(* Logix 5000 project; controller MV vendor 1 type 14 code 217 rev 31.11; software revision 31.00; part 47 of 53 *)
(* tags used below, declared in another part *)
   CWD : CHECKWORD_FLAGS;
   Delphi_Does_Eng_Func : BOOL;
   MV_MV10_CV1 : PlantItem;   // MV10_CV1
   MV_MV11_CV1 : PlantItem;   // MV11_CV1
   MV_MV12_CV1 : PlantItem;   // MV12_CV1
   MV_MV13_CV1 : PlantItem;   // MV13_CV1
   MV_MV14_CV1 : PlantItem;   // MV14_CV1
   MV_MV15_CV1 : PlantItem;   // MV15_CV1
   MV_MV16_CV1 : PlantItem;   // MV16_CV1
   MV_MV17_CV1 : PlantItem;   // MV17_CV1
   MV_MV18_CV1 : PlantItem;   // MV18_CV1
   MV_MV19_CV1 : PlantItem;   // MV19_CV1
   MV_MV1_CV1 : PlantItem;   // MV1_CV1
   MV_MV2_CV1 : PlantItem;   // MV2_CV1
   MV_MV30_CV1 : PlantItem;   // MV30_CV1
   MV_MV31_CV1 : PlantItem;   // MV31_CV1
   MV_MV32_CV1 : PlantItem;   // MV32_CV1
   MV_MV33_CV1 : PlantItem;   // MV33_CV1
   MV_MV34_CV1 : PlantItem;   // MV34_CV1
   MV_MV3_CV1 : PlantItem;   // MV3_CV1
   MV_MV4_CV1 : PlantItem;   // MV4_CV1
   MV_MV5_CV1 : PlantItem;   // MV5_CV1
   MV_MV6_CV1 : PlantItem;   // MV6_CV1
   MV_MV7_CV1 : PlantItem;   // MV7_CV1
   MV_MV8_CV1 : PlantItem;   // MV8_CV1
   MV_MV9_CV1 : PlantItem;   // MV9_CV1
   MV_N255 : DINT[255];   // Old Format Checkwords To Keep Delphi Indicating Status Correctly.
(* MV_Common, continued *)

ROUTINE MV_Old_Checkword_Relaying   (* ladder *)
// Relay New Item Format To Old CW To Keep Delphi Happy Until Full Changeover.
   0: [XIC(Delphi_Does_Eng_Func) [[XIC(MV_N255[0].8) [OTL(MV_MV1_CV1.CW.[CWD.MANUAL]) ,XIC(MV_N255[0].9) OTL(MV_MV1_CV1.CW.[CWD.MANDRV]) ,XIO(MV_N255[0].9) OTU(MV_MV1_CV1.CW.[CWD.MANDRV]) ] ,XIO(MV_N255[0].8) [OTU(MV_MV1_CV1.CW.[CWD.MANUAL]) ,[XIC(MV_MV1_CV1.CW.[CWD.OUTPUT]) OTL(MV_N255[0].9) ,XIO(MV_MV1_CV1.CW.[CWD.OUTPUT]) OTU(MV_N255[0].9) ] ] ] ,[XIC(MV_N255[0].13) OTL(MV_MV1_CV1.CW.[CWD.CHECKOFF]) ,XIO(MV_N255[0].13) OTU(MV_MV1_CV1.CW.[CWD.CHECKOFF]) ] ] ,XIO(Delphi_Does_Eng_Func) [[XIC(MV_MV1_CV1.CW.[CWD.MANUAL]) OTL(MV_N255[0].8) ,XIO(MV_MV1_CV1.CW.[CWD.MANUAL]) OTU(MV_N255[0].8) ] ,[XIC(MV_MV1_CV1.CW.[CWD.CHECKOFF]) OTL(MV_N255[0].13) ,XIO(MV_MV1_CV1.CW.[CWD.CHECKOFF]) OTU(MV_N255[0].13) ] ,[XIC(MV_MV1_CV1.CW.[CWD.OUTPUT]) OTL(MV_N255[0].9) ,XIO(MV_MV1_CV1.CW.[CWD.OUTPUT]) OTU(MV_N255[0].9) ] ] ,XIC(MV_MV1_CV1.CW.[CWD.OUTPUT]) OTE(MV_N255[0].10) ,XIO(MV_MV1_CV1.CW.[CWD.OUTPUT]) OTE(MV_N255[0].11) ,XIC(MV_MV1_CV1.CW.[CWD.FAULT]) OTE(MV_N255[0].15) ];
   1: [XIC(Delphi_Does_Eng_Func) [[XIC(MV_N255[1].8) [OTL(MV_MV2_CV1.CW.[CWD.MANUAL]) ,XIC(MV_N255[1].9) OTL(MV_MV2_CV1.CW.[CWD.MANDRV]) ,XIO(MV_N255[1].9) OTU(MV_MV2_CV1.CW.[CWD.MANDRV]) ] ,XIO(MV_N255[1].8) [OTU(MV_MV2_CV1.CW.[CWD.MANUAL]) ,[XIC(MV_MV2_CV1.CW.[CWD.OUTPUT]) OTL(MV_N255[1].9) ,XIO(MV_MV2_CV1.CW.[CWD.OUTPUT]) OTU(MV_N255[1].9) ] ] ] ,[XIC(MV_N255[1].13) OTL(MV_MV2_CV1.CW.[CWD.CHECKOFF]) ,XIO(MV_N255[1].13) OTU(MV_MV2_CV1.CW.[CWD.CHECKOFF]) ] ] ,XIO(Delphi_Does_Eng_Func) [[XIC(MV_MV2_CV1.CW.[CWD.MANUAL]) OTL(MV_N255[1].8) ,XIO(MV_MV2_CV1.CW.[CWD.MANUAL]) OTU(MV_N255[1].8) ] ,[XIC(MV_MV2_CV1.CW.[CWD.CHECKOFF]) OTL(MV_N255[1].13) ,XIO(MV_MV2_CV1.CW.[CWD.CHECKOFF]) OTU(MV_N255[1].13) ] ,[XIC(MV_MV2_CV1.CW.[CWD.OUTPUT]) OTL(MV_N255[1].9) ,XIO(MV_MV2_CV1.CW.[CWD.OUTPUT]) OTU(MV_N255[1].9) ] ] ,XIC(MV_MV2_CV1.CW.[CWD.OUTPUT]) OTE(MV_N255[1].10) ,XIO(MV_MV2_CV1.CW.[CWD.OUTPUT]) OTE(MV_N255[1].11) ,XIC(MV_MV2_CV1.CW.[CWD.FAULT]) OTE(MV_N255[1].15) ];
   2: [XIC(Delphi_Does_Eng_Func) [[XIC(MV_N255[2].8) [OTL(MV_MV3_CV1.CW.[CWD.MANUAL]) ,XIC(MV_N255[2].9) OTL(MV_MV3_CV1.CW.[CWD.MANDRV]) ,XIO(MV_N255[2].9) OTU(MV_MV3_CV1.CW.[CWD.MANDRV]) ] ,XIO(MV_N255[2].8) [OTU(MV_MV3_CV1.CW.[CWD.MANUAL]) ,[XIC(MV_MV3_CV1.CW.[CWD.OUTPUT]) OTL(MV_N255[2].9) ,XIO(MV_MV3_CV1.CW.[CWD.OUTPUT]) OTU(MV_N255[2].9) ] ] ] ,[XIC(MV_N255[2].13) OTL(MV_MV3_CV1.CW.[CWD.CHECKOFF]) ,XIO(MV_N255[2].13) OTU(MV_MV3_CV1.CW.[CWD.CHECKOFF]) ] ] ,XIO(Delphi_Does_Eng_Func) [[XIC(MV_MV3_CV1.CW.[CWD.MANUAL]) OTL(MV_N255[2].8) ,XIO(MV_MV3_CV1.CW.[CWD.MANUAL]) OTU(MV_N255[2].8) ] ,[XIC(MV_MV3_CV1.CW.[CWD.CHECKOFF]) OTL(MV_N255[2].13) ,XIO(MV_MV3_CV1.CW.[CWD.CHECKOFF]) OTU(MV_N255[2].13) ] ,[XIC(MV_MV3_CV1.CW.[CWD.OUTPUT]) OTL(MV_N255[2].9) ,XIO(MV_MV3_CV1.CW.[CWD.OUTPUT]) OTU(MV_N255[2].9) ] ] ,XIC(MV_MV3_CV1.CW.[CWD.OUTPUT]) OTE(MV_N255[2].10) ,XIO(MV_MV3_CV1.CW.[CWD.OUTPUT]) OTE(MV_N255[2].11) ,XIC(MV_MV3_CV1.CW.[CWD.FAULT]) OTE(MV_N255[2].15) ];
   3: [XIC(Delphi_Does_Eng_Func) [[XIC(MV_N255[3].8) [OTL(MV_MV4_CV1.CW.[CWD.MANUAL]) ,XIC(MV_N255[3].9) OTL(MV_MV4_CV1.CW.[CWD.MANDRV]) ,XIO(MV_N255[3].9) OTU(MV_MV4_CV1.CW.[CWD.MANDRV]) ] ,XIO(MV_N255[3].8) [OTU(MV_MV4_CV1.CW.[CWD.MANUAL]) ,[XIC(MV_MV4_CV1.CW.[CWD.OUTPUT]) OTL(MV_N255[3].9) ,XIO(MV_MV4_CV1.CW.[CWD.OUTPUT]) OTU(MV_N255[3].9) ] ] ] ,[XIC(MV_N255[3].13) OTL(MV_MV4_CV1.CW.[CWD.CHECKOFF]) ,XIO(MV_N255[3].13) OTU(MV_MV4_CV1.CW.[CWD.CHECKOFF]) ] ] ,XIO(Delphi_Does_Eng_Func) [[XIC(MV_MV4_CV1.CW.[CWD.MANUAL]) OTL(MV_N255[3].8) ,XIO(MV_MV4_CV1.CW.[CWD.MANUAL]) OTU(MV_N255[3].8) ] ,[XIC(MV_MV4_CV1.CW.[CWD.CHECKOFF]) OTL(MV_N255[3].13) ,XIO(MV_MV4_CV1.CW.[CWD.CHECKOFF]) OTU(MV_N255[3].13) ] ,[XIC(MV_MV4_CV1.CW.[CWD.OUTPUT]) OTL(MV_N255[3].9) ,XIO(MV_MV4_CV1.CW.[CWD.OUTPUT]) OTU(MV_N255[3].9) ] ] ,XIC(MV_MV4_CV1.CW.[CWD.OUTPUT]) OTE(MV_N255[3].10) ,XIO(MV_MV4_CV1.CW.[CWD.OUTPUT]) OTE(MV_N255[3].11) ,XIC(MV_MV4_CV1.CW.[CWD.FAULT]) OTE(MV_N255[3].15) ];
   4: [XIC(Delphi_Does_Eng_Func) [[XIC(MV_N255[4].8) [OTL(MV_MV5_CV1.CW.[CWD.MANUAL]) ,XIC(MV_N255[4].9) OTL(MV_MV5_CV1.CW.[CWD.MANDRV]) ,XIO(MV_N255[4].9) OTU(MV_MV5_CV1.CW.[CWD.MANDRV]) ] ,XIO(MV_N255[4].8) [OTU(MV_MV5_CV1.CW.[CWD.MANUAL]) ,[XIC(MV_MV5_CV1.CW.[CWD.OUTPUT]) OTL(MV_N255[4].9) ,XIO(MV_MV5_CV1.CW.[CWD.OUTPUT]) OTU(MV_N255[4].9) ] ] ] ,[XIC(MV_N255[4].13) OTL(MV_MV5_CV1.CW.[CWD.CHECKOFF]) ,XIO(MV_N255[4].13) OTU(MV_MV5_CV1.CW.[CWD.CHECKOFF]) ] ] ,XIO(Delphi_Does_Eng_Func) [[XIC(MV_MV5_CV1.CW.[CWD.MANUAL]) OTL(MV_N255[4].8) ,XIO(MV_MV5_CV1.CW.[CWD.MANUAL]) OTU(MV_N255[4].8) ] ,[XIC(MV_MV5_CV1.CW.[CWD.CHECKOFF]) OTL(MV_N255[4].13) ,XIO(MV_MV5_CV1.CW.[CWD.CHECKOFF]) OTU(MV_N255[4].13) ] ,[XIC(MV_MV5_CV1.CW.[CWD.OUTPUT]) OTL(MV_N255[4].9) ,XIO(MV_MV5_CV1.CW.[CWD.OUTPUT]) OTU(MV_N255[4].9) ] ] ,XIC(MV_MV5_CV1.CW.[CWD.OUTPUT]) OTE(MV_N255[4].10) ,XIO(MV_MV5_CV1.CW.[CWD.OUTPUT]) OTE(MV_N255[4].11) ,XIC(MV_MV5_CV1.CW.[CWD.FAULT]) OTE(MV_N255[4].15) ];
   5: [XIC(Delphi_Does_Eng_Func) [[XIC(MV_N255[5].8) [OTL(MV_MV6_CV1.CW.[CWD.MANUAL]) ,XIC(MV_N255[5].9) OTL(MV_MV6_CV1.CW.[CWD.MANDRV]) ,XIO(MV_N255[5].9) OTU(MV_MV6_CV1.CW.[CWD.MANDRV]) ] ,XIO(MV_N255[5].8) [OTU(MV_MV6_CV1.CW.[CWD.MANUAL]) ,[XIC(MV_MV6_CV1.CW.[CWD.OUTPUT]) OTL(MV_N255[5].9) ,XIO(MV_MV6_CV1.CW.[CWD.OUTPUT]) OTU(MV_N255[5].9) ] ] ] ,[XIC(MV_N255[5].13) OTL(MV_MV6_CV1.CW.[CWD.CHECKOFF]) ,XIO(MV_N255[5].13) OTU(MV_MV6_CV1.CW.[CWD.CHECKOFF]) ] ] ,XIO(Delphi_Does_Eng_Func) [[XIC(MV_MV6_CV1.CW.[CWD.MANUAL]) OTL(MV_N255[5].8) ,XIO(MV_MV6_CV1.CW.[CWD.MANUAL]) OTU(MV_N255[5].8) ] ,[XIC(MV_MV6_CV1.CW.[CWD.CHECKOFF]) OTL(MV_N255[5].13) ,XIO(MV_MV6_CV1.CW.[CWD.CHECKOFF]) OTU(MV_N255[5].13) ] ,[XIC(MV_MV6_CV1.CW.[CWD.OUTPUT]) OTL(MV_N255[5].9) ,XIO(MV_MV6_CV1.CW.[CWD.OUTPUT]) OTU(MV_N255[5].9) ] ] ,XIC(MV_MV6_CV1.CW.[CWD.OUTPUT]) OTE(MV_N255[5].10) ,XIO(MV_MV6_CV1.CW.[CWD.OUTPUT]) OTE(MV_N255[5].11) ,XIC(MV_MV6_CV1.CW.[CWD.FAULT]) OTE(MV_N255[5].15) ];
   6: [XIC(Delphi_Does_Eng_Func) [[XIC(MV_N255[6].8) [OTL(MV_MV7_CV1.CW.[CWD.MANUAL]) ,XIC(MV_N255[6].9) OTL(MV_MV7_CV1.CW.[CWD.MANDRV]) ,XIO(MV_N255[6].9) OTU(MV_MV7_CV1.CW.[CWD.MANDRV]) ] ,XIO(MV_N255[6].8) [OTU(MV_MV7_CV1.CW.[CWD.MANUAL]) ,[XIC(MV_MV7_CV1.CW.[CWD.OUTPUT]) OTL(MV_N255[6].9) ,XIO(MV_MV7_CV1.CW.[CWD.OUTPUT]) OTU(MV_N255[6].9) ] ] ] ,[XIC(MV_N255[6].13) OTL(MV_MV7_CV1.CW.[CWD.CHECKOFF]) ,XIO(MV_N255[6].13) OTU(MV_MV7_CV1.CW.[CWD.CHECKOFF]) ] ] ,XIO(Delphi_Does_Eng_Func) [[XIC(MV_MV7_CV1.CW.[CWD.MANUAL]) OTL(MV_N255[6].8) ,XIO(MV_MV7_CV1.CW.[CWD.MANUAL]) OTU(MV_N255[6].8) ] ,[XIC(MV_MV7_CV1.CW.[CWD.CHECKOFF]) OTL(MV_N255[6].13) ,XIO(MV_MV7_CV1.CW.[CWD.CHECKOFF]) OTU(MV_N255[6].13) ] ,[XIC(MV_MV7_CV1.CW.[CWD.OUTPUT]) OTL(MV_N255[6].9) ,XIO(MV_MV7_CV1.CW.[CWD.OUTPUT]) OTU(MV_N255[6].9) ] ] ,XIC(MV_MV7_CV1.CW.[CWD.OUTPUT]) OTE(MV_N255[6].10) ,XIO(MV_MV7_CV1.CW.[CWD.OUTPUT]) OTE(MV_N255[6].11) ,XIC(MV_MV7_CV1.CW.[CWD.FAULT]) OTE(MV_N255[6].15) ];
   7: [XIC(Delphi_Does_Eng_Func) [[XIC(MV_N255[7].8) [OTL(MV_MV8_CV1.CW.[CWD.MANUAL]) ,XIC(MV_N255[7].9) OTL(MV_MV8_CV1.CW.[CWD.MANDRV]) ,XIO(MV_N255[7].9) OTU(MV_MV8_CV1.CW.[CWD.MANDRV]) ] ,XIO(MV_N255[7].8) [OTU(MV_MV8_CV1.CW.[CWD.MANUAL]) ,[XIC(MV_MV8_CV1.CW.[CWD.OUTPUT]) OTL(MV_N255[7].9) ,XIO(MV_MV8_CV1.CW.[CWD.OUTPUT]) OTU(MV_N255[7].9) ] ] ] ,[XIC(MV_N255[7].13) OTL(MV_MV8_CV1.CW.[CWD.CHECKOFF]) ,XIO(MV_N255[7].13) OTU(MV_MV8_CV1.CW.[CWD.CHECKOFF]) ] ] ,XIO(Delphi_Does_Eng_Func) [[XIC(MV_MV8_CV1.CW.[CWD.MANUAL]) OTL(MV_N255[7].8) ,XIO(MV_MV8_CV1.CW.[CWD.MANUAL]) OTU(MV_N255[7].8) ] ,[XIC(MV_MV8_CV1.CW.[CWD.CHECKOFF]) OTL(MV_N255[7].13) ,XIO(MV_MV8_CV1.CW.[CWD.CHECKOFF]) OTU(MV_N255[7].13) ] ,[XIC(MV_MV8_CV1.CW.[CWD.OUTPUT]) OTL(MV_N255[7].9) ,XIO(MV_MV8_CV1.CW.[CWD.OUTPUT]) OTU(MV_N255[7].9) ] ] ,XIC(MV_MV8_CV1.CW.[CWD.OUTPUT]) OTE(MV_N255[7].10) ,XIO(MV_MV8_CV1.CW.[CWD.OUTPUT]) OTE(MV_N255[7].11) ,XIC(MV_MV8_CV1.CW.[CWD.FAULT]) OTE(MV_N255[7].15) ];
   8: [XIC(Delphi_Does_Eng_Func) [[XIC(MV_N255[8].8) [OTL(MV_MV9_CV1.CW.[CWD.MANUAL]) ,XIC(MV_N255[8].9) OTL(MV_MV9_CV1.CW.[CWD.MANDRV]) ,XIO(MV_N255[8].9) OTU(MV_MV9_CV1.CW.[CWD.MANDRV]) ] ,XIO(MV_N255[8].8) [OTU(MV_MV9_CV1.CW.[CWD.MANUAL]) ,[XIC(MV_MV9_CV1.CW.[CWD.OUTPUT]) OTL(MV_N255[8].9) ,XIO(MV_MV9_CV1.CW.[CWD.OUTPUT]) OTU(MV_N255[8].9) ] ] ] ,[XIC(MV_N255[8].13) OTL(MV_MV9_CV1.CW.[CWD.CHECKOFF]) ,XIO(MV_N255[8].13) OTU(MV_MV9_CV1.CW.[CWD.CHECKOFF]) ] ] ,XIO(Delphi_Does_Eng_Func) [[XIC(MV_MV9_CV1.CW.[CWD.MANUAL]) OTL(MV_N255[8].8) ,XIO(MV_MV9_CV1.CW.[CWD.MANUAL]) OTU(MV_N255[8].8) ] ,[XIC(MV_MV9_CV1.CW.[CWD.CHECKOFF]) OTL(MV_N255[8].13) ,XIO(MV_MV9_CV1.CW.[CWD.CHECKOFF]) OTU(MV_N255[8].13) ] ,[XIC(MV_MV9_CV1.CW.[CWD.OUTPUT]) OTL(MV_N255[8].9) ,XIO(MV_MV9_CV1.CW.[CWD.OUTPUT]) OTU(MV_N255[8].9) ] ] ,XIC(MV_MV9_CV1.CW.[CWD.OUTPUT]) OTE(MV_N255[8].10) ,XIO(MV_MV9_CV1.CW.[CWD.OUTPUT]) OTE(MV_N255[8].11) ,XIC(MV_MV9_CV1.CW.[CWD.FAULT]) OTE(MV_N255[8].15) ];
   9: [XIC(Delphi_Does_Eng_Func) [[XIC(MV_N255[9].8) [OTL(MV_MV10_CV1.CW.[CWD.MANUAL]) ,XIC(MV_N255[9].9) OTL(MV_MV10_CV1.CW.[CWD.MANDRV]) ,XIO(MV_N255[9].9) OTU(MV_MV10_CV1.CW.[CWD.MANDRV]) ] ,XIO(MV_N255[9].8) [OTU(MV_MV10_CV1.CW.[CWD.MANUAL]) ,[XIC(MV_MV10_CV1.CW.[CWD.OUTPUT]) OTL(MV_N255[9].9) ,XIO(MV_MV10_CV1.CW.[CWD.OUTPUT]) OTU(MV_N255[9].9) ] ] ] ,[XIC(MV_N255[9].13) OTL(MV_MV10_CV1.CW.[CWD.CHECKOFF]) ,XIO(MV_N255[9].13) OTU(MV_MV10_CV1.CW.[CWD.CHECKOFF]) ] ] ,XIO(Delphi_Does_Eng_Func) [[XIC(MV_MV10_CV1.CW.[CWD.MANUAL]) OTL(MV_N255[9].8) ,XIO(MV_MV10_CV1.CW.[CWD.MANUAL]) OTU(MV_N255[9].8) ] ,[XIC(MV_MV10_CV1.CW.[CWD.CHECKOFF]) OTL(MV_N255[9].13) ,XIO(MV_MV10_CV1.CW.[CWD.CHECKOFF]) OTU(MV_N255[9].13) ] ,[XIC(MV_MV10_CV1.CW.[CWD.OUTPUT]) OTL(MV_N255[9].9) ,XIO(MV_MV10_CV1.CW.[CWD.OUTPUT]) OTU(MV_N255[9].9) ] ] ,XIC(MV_MV10_CV1.CW.[CWD.OUTPUT]) OTE(MV_N255[9].10) ,XIO(MV_MV10_CV1.CW.[CWD.OUTPUT]) OTE(MV_N255[9].11) ,XIC(MV_MV10_CV1.CW.[CWD.FAULT]) OTE(MV_N255[9].15) ];
   10: [XIC(Delphi_Does_Eng_Func) [[XIC(MV_N255[10].8) [OTL(MV_MV11_CV1.CW.[CWD.MANUAL]) ,XIC(MV_N255[10].9) OTL(MV_MV11_CV1.CW.[CWD.MANDRV]) ,XIO(MV_N255[10].9) OTU(MV_MV11_CV1.CW.[CWD.MANDRV]) ] ,XIO(MV_N255[10].8) [OTU(MV_MV11_CV1.CW.[CWD.MANUAL]) ,[XIC(MV_MV11_CV1.CW.[CWD.OUTPUT]) OTL(MV_N255[10].9) ,XIO(MV_MV11_CV1.CW.[CWD.OUTPUT]) OTU(MV_N255[10].9) ] ] ] ,[XIC(MV_N255[10].13) OTL(MV_MV11_CV1.CW.[CWD.CHECKOFF]) ,XIO(MV_N255[10].13) OTU(MV_MV11_CV1.CW.[CWD.CHECKOFF]) ] ] ,XIO(Delphi_Does_Eng_Func) [[XIC(MV_MV11_CV1.CW.[CWD.MANUAL]) OTL(MV_N255[10].8) ,XIO(MV_MV11_CV1.CW.[CWD.MANUAL]) OTU(MV_N255[10].8) ] ,[XIC(MV_MV11_CV1.CW.[CWD.CHECKOFF]) OTL(MV_N255[10].13) ,XIO(MV_MV11_CV1.CW.[CWD.CHECKOFF]) OTU(MV_N255[10].13) ] ,[XIC(MV_MV11_CV1.CW.[CWD.OUTPUT]) OTL(MV_N255[10].9) ,XIO(MV_MV11_CV1.CW.[CWD.OUTPUT]) OTU(MV_N255[10].9) ] ] ,XIC(MV_MV11_CV1.CW.[CWD.OUTPUT]) OTE(MV_N255[10].10) ,XIO(MV_MV11_CV1.CW.[CWD.OUTPUT]) OTE(MV_N255[10].11) ,XIC(MV_MV11_CV1.CW.[CWD.FAULT]) OTE(MV_N255[10].15) ];
   11: [XIC(Delphi_Does_Eng_Func) [[XIC(MV_N255[11].8) [OTL(MV_MV12_CV1.CW.[CWD.MANUAL]) ,XIC(MV_N255[11].9) OTL(MV_MV12_CV1.CW.[CWD.MANDRV]) ,XIO(MV_N255[11].9) OTU(MV_MV12_CV1.CW.[CWD.MANDRV]) ] ,XIO(MV_N255[11].8) [OTU(MV_MV12_CV1.CW.[CWD.MANUAL]) ,[XIC(MV_MV12_CV1.CW.[CWD.OUTPUT]) OTL(MV_N255[11].9) ,XIO(MV_MV12_CV1.CW.[CWD.OUTPUT]) OTU(MV_N255[11].9) ] ] ] ,[XIC(MV_N255[11].13) OTL(MV_MV12_CV1.CW.[CWD.CHECKOFF]) ,XIO(MV_N255[11].13) OTU(MV_MV12_CV1.CW.[CWD.CHECKOFF]) ] ] ,XIO(Delphi_Does_Eng_Func) [[XIC(MV_MV12_CV1.CW.[CWD.MANUAL]) OTL(MV_N255[11].8) ,XIO(MV_MV12_CV1.CW.[CWD.MANUAL]) OTU(MV_N255[11].8) ] ,[XIC(MV_MV12_CV1.CW.[CWD.CHECKOFF]) OTL(MV_N255[11].13) ,XIO(MV_MV12_CV1.CW.[CWD.CHECKOFF]) OTU(MV_N255[11].13) ] ,[XIC(MV_MV12_CV1.CW.[CWD.OUTPUT]) OTL(MV_N255[11].9) ,XIO(MV_MV12_CV1.CW.[CWD.OUTPUT]) OTU(MV_N255[11].9) ] ] ,XIC(MV_MV12_CV1.CW.[CWD.OUTPUT]) OTE(MV_N255[11].10) ,XIO(MV_MV12_CV1.CW.[CWD.OUTPUT]) OTE(MV_N255[11].11) ,XIC(MV_MV12_CV1.CW.[CWD.FAULT]) OTE(MV_N255[11].15) ];
   12: [XIC(Delphi_Does_Eng_Func) [[XIC(MV_N255[12].8) [OTL(MV_MV13_CV1.CW.[CWD.MANUAL]) ,XIC(MV_N255[12].9) OTL(MV_MV13_CV1.CW.[CWD.MANDRV]) ,XIO(MV_N255[12].9) OTU(MV_MV13_CV1.CW.[CWD.MANDRV]) ] ,XIO(MV_N255[12].8) [OTU(MV_MV13_CV1.CW.[CWD.MANUAL]) ,[XIC(MV_MV13_CV1.CW.[CWD.OUTPUT]) OTL(MV_N255[12].9) ,XIO(MV_MV13_CV1.CW.[CWD.OUTPUT]) OTU(MV_N255[12].9) ] ] ] ,[XIC(MV_N255[12].13) OTL(MV_MV13_CV1.CW.[CWD.CHECKOFF]) ,XIO(MV_N255[12].13) OTU(MV_MV13_CV1.CW.[CWD.CHECKOFF]) ] ] ,XIO(Delphi_Does_Eng_Func) [[XIC(MV_MV13_CV1.CW.[CWD.MANUAL]) OTL(MV_N255[12].8) ,XIO(MV_MV13_CV1.CW.[CWD.MANUAL]) OTU(MV_N255[12].8) ] ,[XIC(MV_MV13_CV1.CW.[CWD.CHECKOFF]) OTL(MV_N255[12].13) ,XIO(MV_MV13_CV1.CW.[CWD.CHECKOFF]) OTU(MV_N255[12].13) ] ,[XIC(MV_MV13_CV1.CW.[CWD.OUTPUT]) OTL(MV_N255[12].9) ,XIO(MV_MV13_CV1.CW.[CWD.OUTPUT]) OTU(MV_N255[12].9) ] ] ,XIC(MV_MV13_CV1.CW.[CWD.OUTPUT]) OTE(MV_N255[12].10) ,XIO(MV_MV13_CV1.CW.[CWD.OUTPUT]) OTE(MV_N255[12].11) ,XIC(MV_MV13_CV1.CW.[CWD.FAULT]) OTE(MV_N255[12].15) ];
   13: [XIC(Delphi_Does_Eng_Func) [[XIC(MV_N255[13].8) [OTL(MV_MV14_CV1.CW.[CWD.MANUAL]) ,XIC(MV_N255[13].9) OTL(MV_MV14_CV1.CW.[CWD.MANDRV]) ,XIO(MV_N255[13].9) OTU(MV_MV14_CV1.CW.[CWD.MANDRV]) ] ,XIO(MV_N255[13].8) [OTU(MV_MV14_CV1.CW.[CWD.MANUAL]) ,[XIC(MV_MV14_CV1.CW.[CWD.OUTPUT]) OTL(MV_N255[13].9) ,XIO(MV_MV14_CV1.CW.[CWD.OUTPUT]) OTU(MV_N255[13].9) ] ] ] ,[XIC(MV_N255[13].13) OTL(MV_MV14_CV1.CW.[CWD.CHECKOFF]) ,XIO(MV_N255[13].13) OTU(MV_MV14_CV1.CW.[CWD.CHECKOFF]) ] ] ,XIO(Delphi_Does_Eng_Func) [[XIC(MV_MV14_CV1.CW.[CWD.MANUAL]) OTL(MV_N255[13].8) ,XIO(MV_MV14_CV1.CW.[CWD.MANUAL]) OTU(MV_N255[13].8) ] ,[XIC(MV_MV14_CV1.CW.[CWD.CHECKOFF]) OTL(MV_N255[13].13) ,XIO(MV_MV14_CV1.CW.[CWD.CHECKOFF]) OTU(MV_N255[13].13) ] ,[XIC(MV_MV14_CV1.CW.[CWD.OUTPUT]) OTL(MV_N255[13].9) ,XIO(MV_MV14_CV1.CW.[CWD.OUTPUT]) OTU(MV_N255[13].9) ] ] ,XIC(MV_MV14_CV1.CW.[CWD.OUTPUT]) OTE(MV_N255[13].10) ,XIO(MV_MV14_CV1.CW.[CWD.OUTPUT]) OTE(MV_N255[13].11) ,XIC(MV_MV14_CV1.CW.[CWD.FAULT]) OTE(MV_N255[13].15) ];
   14: [XIC(Delphi_Does_Eng_Func) [[XIC(MV_N255[14].8) [OTL(MV_MV15_CV1.CW.[CWD.MANUAL]) ,XIC(MV_N255[14].9) OTL(MV_MV15_CV1.CW.[CWD.MANDRV]) ,XIO(MV_N255[14].9) OTU(MV_MV15_CV1.CW.[CWD.MANDRV]) ] ,XIO(MV_N255[14].8) [OTU(MV_MV15_CV1.CW.[CWD.MANUAL]) ,[XIC(MV_MV15_CV1.CW.[CWD.OUTPUT]) OTL(MV_N255[14].9) ,XIO(MV_MV15_CV1.CW.[CWD.OUTPUT]) OTU(MV_N255[14].9) ] ] ] ,[XIC(MV_N255[14].13) OTL(MV_MV15_CV1.CW.[CWD.CHECKOFF]) ,XIO(MV_N255[14].13) OTU(MV_MV15_CV1.CW.[CWD.CHECKOFF]) ] ] ,XIO(Delphi_Does_Eng_Func) [[XIC(MV_MV15_CV1.CW.[CWD.MANUAL]) OTL(MV_N255[14].8) ,XIO(MV_MV15_CV1.CW.[CWD.MANUAL]) OTU(MV_N255[14].8) ] ,[XIC(MV_MV15_CV1.CW.[CWD.CHECKOFF]) OTL(MV_N255[14].13) ,XIO(MV_MV15_CV1.CW.[CWD.CHECKOFF]) OTU(MV_N255[14].13) ] ,[XIC(MV_MV15_CV1.CW.[CWD.OUTPUT]) OTL(MV_N255[14].9) ,XIO(MV_MV15_CV1.CW.[CWD.OUTPUT]) OTU(MV_N255[14].9) ] ] ,XIC(MV_MV15_CV1.CW.[CWD.OUTPUT]) OTE(MV_N255[14].10) ,XIO(MV_MV15_CV1.CW.[CWD.OUTPUT]) OTE(MV_N255[14].11) ,XIC(MV_MV15_CV1.CW.[CWD.FAULT]) OTE(MV_N255[14].15) ];
   15: [XIC(Delphi_Does_Eng_Func) [[XIC(MV_N255[15].8) [OTL(MV_MV16_CV1.CW.[CWD.MANUAL]) ,XIC(MV_N255[15].9) OTL(MV_MV16_CV1.CW.[CWD.MANDRV]) ,XIO(MV_N255[15].9) OTU(MV_MV16_CV1.CW.[CWD.MANDRV]) ] ,XIO(MV_N255[15].8) [OTU(MV_MV16_CV1.CW.[CWD.MANUAL]) ,[XIC(MV_MV16_CV1.CW.[CWD.OUTPUT]) OTL(MV_N255[15].9) ,XIO(MV_MV16_CV1.CW.[CWD.OUTPUT]) OTU(MV_N255[15].9) ] ] ] ,[XIC(MV_N255[15].13) OTL(MV_MV16_CV1.CW.[CWD.CHECKOFF]) ,XIO(MV_N255[15].13) OTU(MV_MV16_CV1.CW.[CWD.CHECKOFF]) ] ] ,XIO(Delphi_Does_Eng_Func) [[XIC(MV_MV16_CV1.CW.[CWD.MANUAL]) OTL(MV_N255[15].8) ,XIO(MV_MV16_CV1.CW.[CWD.MANUAL]) OTU(MV_N255[15].8) ] ,[XIC(MV_MV16_CV1.CW.[CWD.CHECKOFF]) OTL(MV_N255[15].13) ,XIO(MV_MV16_CV1.CW.[CWD.CHECKOFF]) OTU(MV_N255[15].13) ] ,[XIC(MV_MV16_CV1.CW.[CWD.OUTPUT]) OTL(MV_N255[15].9) ,XIO(MV_MV16_CV1.CW.[CWD.OUTPUT]) OTU(MV_N255[15].9) ] ] ,XIC(MV_MV16_CV1.CW.[CWD.OUTPUT]) OTE(MV_N255[15].10) ,XIO(MV_MV16_CV1.CW.[CWD.OUTPUT]) OTE(MV_N255[15].11) ,XIC(MV_MV16_CV1.CW.[CWD.FAULT]) OTE(MV_N255[15].15) ];
   16: [XIC(Delphi_Does_Eng_Func) [[XIC(MV_N255[16].8) [OTL(MV_MV17_CV1.CW.[CWD.MANUAL]) ,XIC(MV_N255[16].9) OTL(MV_MV17_CV1.CW.[CWD.MANDRV]) ,XIO(MV_N255[16].9) OTU(MV_MV17_CV1.CW.[CWD.MANDRV]) ] ,XIO(MV_N255[16].8) [OTU(MV_MV17_CV1.CW.[CWD.MANUAL]) ,[XIC(MV_MV17_CV1.CW.[CWD.OUTPUT]) OTL(MV_N255[16].9) ,XIO(MV_MV17_CV1.CW.[CWD.OUTPUT]) OTU(MV_N255[16].9) ] ] ] ,[XIC(MV_N255[16].13) OTL(MV_MV17_CV1.CW.[CWD.CHECKOFF]) ,XIO(MV_N255[16].13) OTU(MV_MV17_CV1.CW.[CWD.CHECKOFF]) ] ] ,XIO(Delphi_Does_Eng_Func) [[XIC(MV_MV17_CV1.CW.[CWD.MANUAL]) OTL(MV_N255[16].8) ,XIO(MV_MV17_CV1.CW.[CWD.MANUAL]) OTU(MV_N255[16].8) ] ,[XIC(MV_MV17_CV1.CW.[CWD.CHECKOFF]) OTL(MV_N255[16].13) ,XIO(MV_MV17_CV1.CW.[CWD.CHECKOFF]) OTU(MV_N255[16].13) ] ,[XIC(MV_MV17_CV1.CW.[CWD.OUTPUT]) OTL(MV_N255[16].9) ,XIO(MV_MV17_CV1.CW.[CWD.OUTPUT]) OTU(MV_N255[16].9) ] ] ,XIC(MV_MV17_CV1.CW.[CWD.OUTPUT]) OTE(MV_N255[16].10) ,XIO(MV_MV17_CV1.CW.[CWD.OUTPUT]) OTE(MV_N255[16].11) ,XIC(MV_MV17_CV1.CW.[CWD.FAULT]) OTE(MV_N255[16].15) ];
   17: [XIC(Delphi_Does_Eng_Func) [[XIC(MV_N255[17].8) [OTL(MV_MV18_CV1.CW.[CWD.MANUAL]) ,XIC(MV_N255[17].9) OTL(MV_MV18_CV1.CW.[CWD.MANDRV]) ,XIO(MV_N255[17].9) OTU(MV_MV18_CV1.CW.[CWD.MANDRV]) ] ,XIO(MV_N255[17].8) [OTU(MV_MV18_CV1.CW.[CWD.MANUAL]) ,[XIC(MV_MV18_CV1.CW.[CWD.OUTPUT]) OTL(MV_N255[17].9) ,XIO(MV_MV18_CV1.CW.[CWD.OUTPUT]) OTU(MV_N255[17].9) ] ] ] ,[XIC(MV_N255[17].13) OTL(MV_MV18_CV1.CW.[CWD.CHECKOFF]) ,XIO(MV_N255[17].13) OTU(MV_MV18_CV1.CW.[CWD.CHECKOFF]) ] ] ,XIO(Delphi_Does_Eng_Func) [[XIC(MV_MV18_CV1.CW.[CWD.MANUAL]) OTL(MV_N255[17].8) ,XIO(MV_MV18_CV1.CW.[CWD.MANUAL]) OTU(MV_N255[17].8) ] ,[XIC(MV_MV18_CV1.CW.[CWD.CHECKOFF]) OTL(MV_N255[17].13) ,XIO(MV_MV18_CV1.CW.[CWD.CHECKOFF]) OTU(MV_N255[17].13) ] ,[XIC(MV_MV18_CV1.CW.[CWD.OUTPUT]) OTL(MV_N255[17].9) ,XIO(MV_MV18_CV1.CW.[CWD.OUTPUT]) OTU(MV_N255[17].9) ] ] ,XIC(MV_MV18_CV1.CW.[CWD.OUTPUT]) OTE(MV_N255[17].10) ,XIO(MV_MV18_CV1.CW.[CWD.OUTPUT]) OTE(MV_N255[17].11) ,XIC(MV_MV18_CV1.CW.[CWD.FAULT]) OTE(MV_N255[17].15) ];
   18: [XIC(Delphi_Does_Eng_Func) [[XIC(MV_N255[18].8) [OTL(MV_MV19_CV1.CW.[CWD.MANUAL]) ,XIC(MV_N255[18].9) OTL(MV_MV19_CV1.CW.[CWD.MANDRV]) ,XIO(MV_N255[18].9) OTU(MV_MV19_CV1.CW.[CWD.MANDRV]) ] ,XIO(MV_N255[18].8) [OTU(MV_MV19_CV1.CW.[CWD.MANUAL]) ,[XIC(MV_MV19_CV1.CW.[CWD.OUTPUT]) OTL(MV_N255[18].9) ,XIO(MV_MV19_CV1.CW.[CWD.OUTPUT]) OTU(MV_N255[18].9) ] ] ] ,[XIC(MV_N255[18].13) OTL(MV_MV19_CV1.CW.[CWD.CHECKOFF]) ,XIO(MV_N255[18].13) OTU(MV_MV19_CV1.CW.[CWD.CHECKOFF]) ] ] ,XIO(Delphi_Does_Eng_Func) [[XIC(MV_MV19_CV1.CW.[CWD.MANUAL]) OTL(MV_N255[18].8) ,XIO(MV_MV19_CV1.CW.[CWD.MANUAL]) OTU(MV_N255[18].8) ] ,[XIC(MV_MV19_CV1.CW.[CWD.CHECKOFF]) OTL(MV_N255[18].13) ,XIO(MV_MV19_CV1.CW.[CWD.CHECKOFF]) OTU(MV_N255[18].13) ] ,[XIC(MV_MV19_CV1.CW.[CWD.OUTPUT]) OTL(MV_N255[18].9) ,XIO(MV_MV19_CV1.CW.[CWD.OUTPUT]) OTU(MV_N255[18].9) ] ] ,XIC(MV_MV19_CV1.CW.[CWD.OUTPUT]) OTE(MV_N255[18].10) ,XIO(MV_MV19_CV1.CW.[CWD.OUTPUT]) OTE(MV_N255[18].11) ,XIC(MV_MV19_CV1.CW.[CWD.FAULT]) OTE(MV_N255[18].15) ];
   19: [XIC(Delphi_Does_Eng_Func) [[XIC(MV_N255[19].8) [OTL(MV_MV30_CV1.CW.[CWD.MANUAL]) ,XIC(MV_N255[19].9) OTL(MV_MV30_CV1.CW.[CWD.MANDRV]) ,XIO(MV_N255[19].9) OTU(MV_MV30_CV1.CW.[CWD.MANDRV]) ] ,XIO(MV_N255[19].8) [OTU(MV_MV30_CV1.CW.[CWD.MANUAL]) ,[XIC(MV_MV30_CV1.CW.[CWD.OUTPUT]) OTL(MV_N255[19].9) ,XIO(MV_MV30_CV1.CW.[CWD.OUTPUT]) OTU(MV_N255[19].9) ] ] ] ,[XIC(MV_N255[19].13) OTL(MV_MV30_CV1.CW.[CWD.CHECKOFF]) ,XIO(MV_N255[19].13) OTU(MV_MV30_CV1.CW.[CWD.CHECKOFF]) ] ] ,XIO(Delphi_Does_Eng_Func) [[XIC(MV_MV30_CV1.CW.[CWD.MANUAL]) OTL(MV_N255[19].8) ,XIO(MV_MV30_CV1.CW.[CWD.MANUAL]) OTU(MV_N255[19].8) ] ,[XIC(MV_MV30_CV1.CW.[CWD.CHECKOFF]) OTL(MV_N255[19].13) ,XIO(MV_MV30_CV1.CW.[CWD.CHECKOFF]) OTU(MV_N255[19].13) ] ,[XIC(MV_MV30_CV1.CW.[CWD.OUTPUT]) OTL(MV_N255[19].9) ,XIO(MV_MV30_CV1.CW.[CWD.OUTPUT]) OTU(MV_N255[19].9) ] ] ,XIC(MV_MV30_CV1.CW.[CWD.OUTPUT]) OTE(MV_N255[19].10) ,XIO(MV_MV30_CV1.CW.[CWD.OUTPUT]) OTE(MV_N255[19].11) ,XIC(MV_MV30_CV1.CW.[CWD.FAULT]) OTE(MV_N255[19].15) ];
   20: [XIC(Delphi_Does_Eng_Func) [[XIC(MV_N255[20].8) [OTL(MV_MV31_CV1.CW.[CWD.MANUAL]) ,XIC(MV_N255[20].9) OTL(MV_MV31_CV1.CW.[CWD.MANDRV]) ,XIO(MV_N255[20].9) OTU(MV_MV31_CV1.CW.[CWD.MANDRV]) ] ,XIO(MV_N255[20].8) [OTU(MV_MV31_CV1.CW.[CWD.MANUAL]) ,[XIC(MV_MV31_CV1.CW.[CWD.OUTPUT]) OTL(MV_N255[20].9) ,XIO(MV_MV31_CV1.CW.[CWD.OUTPUT]) OTU(MV_N255[20].9) ] ] ] ,[XIC(MV_N255[20].13) OTL(MV_MV31_CV1.CW.[CWD.CHECKOFF]) ,XIO(MV_N255[20].13) OTU(MV_MV31_CV1.CW.[CWD.CHECKOFF]) ] ] ,XIO(Delphi_Does_Eng_Func) [[XIC(MV_MV31_CV1.CW.[CWD.MANUAL]) OTL(MV_N255[20].8) ,XIO(MV_MV31_CV1.CW.[CWD.MANUAL]) OTU(MV_N255[20].8) ] ,[XIC(MV_MV31_CV1.CW.[CWD.CHECKOFF]) OTL(MV_N255[20].13) ,XIO(MV_MV31_CV1.CW.[CWD.CHECKOFF]) OTU(MV_N255[20].13) ] ,[XIC(MV_MV31_CV1.CW.[CWD.OUTPUT]) OTL(MV_N255[20].9) ,XIO(MV_MV31_CV1.CW.[CWD.OUTPUT]) OTU(MV_N255[20].9) ] ] ,XIC(MV_MV31_CV1.CW.[CWD.OUTPUT]) OTE(MV_N255[20].10) ,XIO(MV_MV31_CV1.CW.[CWD.OUTPUT]) OTE(MV_N255[20].11) ,XIC(MV_MV31_CV1.CW.[CWD.FAULT]) OTE(MV_N255[20].15) ];
   21: [XIC(Delphi_Does_Eng_Func) [[XIC(MV_N255[21].8) [OTL(MV_MV32_CV1.CW.[CWD.MANUAL]) ,XIC(MV_N255[21].9) OTL(MV_MV32_CV1.CW.[CWD.MANDRV]) ,XIO(MV_N255[21].9) OTU(MV_MV32_CV1.CW.[CWD.MANDRV]) ] ,XIO(MV_N255[21].8) [OTU(MV_MV32_CV1.CW.[CWD.MANUAL]) ,[XIC(MV_MV32_CV1.CW.[CWD.OUTPUT]) OTL(MV_N255[21].9) ,XIO(MV_MV32_CV1.CW.[CWD.OUTPUT]) OTU(MV_N255[21].9) ] ] ] ,[XIC(MV_N255[21].13) OTL(MV_MV32_CV1.CW.[CWD.CHECKOFF]) ,XIO(MV_N255[21].13) OTU(MV_MV32_CV1.CW.[CWD.CHECKOFF]) ] ] ,XIO(Delphi_Does_Eng_Func) [[XIC(MV_MV32_CV1.CW.[CWD.MANUAL]) OTL(MV_N255[21].8) ,XIO(MV_MV32_CV1.CW.[CWD.MANUAL]) OTU(MV_N255[21].8) ] ,[XIC(MV_MV32_CV1.CW.[CWD.CHECKOFF]) OTL(MV_N255[21].13) ,XIO(MV_MV32_CV1.CW.[CWD.CHECKOFF]) OTU(MV_N255[21].13) ] ,[XIC(MV_MV32_CV1.CW.[CWD.OUTPUT]) OTL(MV_N255[21].9) ,XIO(MV_MV32_CV1.CW.[CWD.OUTPUT]) OTU(MV_N255[21].9) ] ] ,XIC(MV_MV32_CV1.CW.[CWD.OUTPUT]) OTE(MV_N255[21].10) ,XIO(MV_MV32_CV1.CW.[CWD.OUTPUT]) OTE(MV_N255[21].11) ,XIC(MV_MV32_CV1.CW.[CWD.FAULT]) OTE(MV_N255[21].15) ];
   22: [XIC(Delphi_Does_Eng_Func) [[XIC(MV_N255[22].8) [OTL(MV_MV33_CV1.CW.[CWD.MANUAL]) ,XIC(MV_N255[22].9) OTL(MV_MV33_CV1.CW.[CWD.MANDRV]) ,XIO(MV_N255[22].9) OTU(MV_MV33_CV1.CW.[CWD.MANDRV]) ] ,XIO(MV_N255[22].8) [OTU(MV_MV33_CV1.CW.[CWD.MANUAL]) ,[XIC(MV_MV33_CV1.CW.[CWD.OUTPUT]) OTL(MV_N255[22].9) ,XIO(MV_MV33_CV1.CW.[CWD.OUTPUT]) OTU(MV_N255[22].9) ] ] ] ,[XIC(MV_N255[22].13) OTL(MV_MV33_CV1.CW.[CWD.CHECKOFF]) ,XIO(MV_N255[22].13) OTU(MV_MV33_CV1.CW.[CWD.CHECKOFF]) ] ] ,XIO(Delphi_Does_Eng_Func) [[XIC(MV_MV33_CV1.CW.[CWD.MANUAL]) OTL(MV_N255[22].8) ,XIO(MV_MV33_CV1.CW.[CWD.MANUAL]) OTU(MV_N255[22].8) ] ,[XIC(MV_MV33_CV1.CW.[CWD.CHECKOFF]) OTL(MV_N255[22].13) ,XIO(MV_MV33_CV1.CW.[CWD.CHECKOFF]) OTU(MV_N255[22].13) ] ,[XIC(MV_MV33_CV1.CW.[CWD.OUTPUT]) OTL(MV_N255[22].9) ,XIO(MV_MV33_CV1.CW.[CWD.OUTPUT]) OTU(MV_N255[22].9) ] ] ,XIC(MV_MV33_CV1.CW.[CWD.OUTPUT]) OTE(MV_N255[22].10) ,XIO(MV_MV33_CV1.CW.[CWD.OUTPUT]) OTE(MV_N255[22].11) ,XIC(MV_MV33_CV1.CW.[CWD.FAULT]) OTE(MV_N255[22].15) ];
   23: [XIC(Delphi_Does_Eng_Func) [[XIC(MV_N255[23].8) [OTL(MV_MV34_CV1.CW.[CWD.MANUAL]) ,XIC(MV_N255[23].9) OTL(MV_MV34_CV1.CW.[CWD.MANDRV]) ,XIO(MV_N255[23].9) OTU(MV_MV34_CV1.CW.[CWD.MANDRV]) ] ,XIO(MV_N255[23].8) [OTU(MV_MV34_CV1.CW.[CWD.MANUAL]) ,[XIC(MV_MV34_CV1.CW.[CWD.OUTPUT]) OTL(MV_N255[23].9) ,XIO(MV_MV34_CV1.CW.[CWD.OUTPUT]) OTU(MV_N255[23].9) ] ] ] ,[XIC(MV_N255[23].13) OTL(MV_MV34_CV1.CW.[CWD.CHECKOFF]) ,XIO(MV_N255[23].13) OTU(MV_MV34_CV1.CW.[CWD.CHECKOFF]) ] ] ,XIO(Delphi_Does_Eng_Func) [[XIC(MV_MV34_CV1.CW.[CWD.MANUAL]) OTL(MV_N255[23].8) ,XIO(MV_MV34_CV1.CW.[CWD.MANUAL]) OTU(MV_N255[23].8) ] ,[XIC(MV_MV34_CV1.CW.[CWD.CHECKOFF]) OTL(MV_N255[23].13) ,XIO(MV_MV34_CV1.CW.[CWD.CHECKOFF]) OTU(MV_N255[23].13) ] ,[XIC(MV_MV34_CV1.CW.[CWD.OUTPUT]) OTL(MV_N255[23].9) ,XIO(MV_MV34_CV1.CW.[CWD.OUTPUT]) OTU(MV_N255[23].9) ] ] ,XIC(MV_MV34_CV1.CW.[CWD.OUTPUT]) OTE(MV_N255[23].10) ,XIO(MV_MV34_CV1.CW.[CWD.OUTPUT]) OTE(MV_N255[23].11) ,XIC(MV_MV34_CV1.CW.[CWD.FAULT]) OTE(MV_N255[23].15) ];
